// TIA Portal project "EMS" (V15.1)

(* hardware
DEVICE "HMI_SDC"  TP1500 Comfort
   slot 0: "HMI_SDC"  TP1500 Comfort  6AV2 124-0QC02-0AX1  15.1.0.0
   slot 1: "HMI_RT_2"  TP1500 Comfort  6AV2 124-0QC02-0AX1  15.1.0.0
   slot 5: "HMI_SDC._CP_2"  PROFINET Interface  15.0.1.0
      slot 1: "PROFINET Schnittstelle_1"  PROFINET Interface
         slot 1: "Port_1"  Port
         slot 2: "Port_2"  Port
   slot 6: "HMI_SDC._CP_1"  PROFINET Interface  15.0.1.0
      slot 1: "PROFINET Schnittstelle_GBit"  PROFINET Interface
         slot 1: "Port_1"  Port
   slot 7: "HMI_SDC.I/DP_CP_1"  MPI/DP Interface  15.0.1.0
DEVICE "SCALANCE W client"  SCALANCE W-Station
   slot 0: "SCALANCE W rack"  Rail
   slot 0: "_wlan"  SCALANCE W734-1 RJ45 US  6GK5 734-1FX00-0AB0  V6.2
DEVICE "S71500/ET200MP station_1"  S7-1500 station
   slot 0: "Rail_0"  Rack  6ES7 590-1***0-0AA0
   slot 1: "SDC_PLC"  CPU 1518F-4 PN/DP  6ES7 518-4FP00-0AB0  V2.6
      slot 3: "CPU display_1"  6ES7591-1BA00-0AA0
   slot 2: "DI 16x24VDC BA_1"  DI 16x24VDC BA  6ES7 521-1BH10-0AA0  V1.0
   slot 3: "DQ 16x24VDC/0.5A BA_1"  DQ 16x24VDC/0.5A BA  6ES7 522-1BH10-0AA0  V1.0
DEVICE "ET 200SP station_2"  ET 200SP-Station
   slot 0: "Rack_0"  Rack  6ES5 710-8MAx1
   slot 1: "_PLC"  CPU 1512SP F-1 PN  6ES7 512-1SK01-0AB0  V2.1
   slot 2: "F-DI 8x24VDC HF_1"  F-DI 8x24VDC HF  6ES7 136-6BA00-0CA0  V1.0
      slot 1: "F-DI 8x24VDC HF_1"  F-DI 8x24VDC HF
   slot 3: "F-DQ 4x24VDC/2A PM HF_1"  F-DQ 4x24VDC/2A PM HF  6ES7 136-6DB00-0CA0  V1.0
      slot 1: "F-DQ 4x24VDC/2A PM HF_1"  F-DQ 4x24VDC/2A PM HF
   slot 4: "DI 16x24VDC ST_1"  DI 16x24VDC ST  6ES7 131-6BH00-0BA0  V1.1
      slot 1: "DI 16x24VDC ST_1"  DI 16x24VDC ST
   slot 5: "DQ 8x24VDC/0.5A ST_1"  DQ 8x24VDC/0.5A ST  6ES7 132-6BF01-0BA0  V0.0
      slot 1: "DQ 8x24VDC/0.5A ST_1"  DQ 8x24VDC/0.5A ST
   slot 6: "Server module_1"  Server module  6ES7 193-6PA00-0AA0  V1.1
      slot 1: "Server module_1"  Server module
   slot 127: "BA 2xRJ45"  BA 2xRJ45  6ES7 193-6AR00-0AA0  V0.0
      slot 32769: "Port_1"  6ES7 193-6AR00-0AA0
      slot 32770: "Port_2"  6ES7 193-6AR00-0AA0
DEVICE "GSD device_4"  GSD.Device.PN
   slot 0: "Rack"  Rack  V1.0
   slot 0: "_DRIVE"  SINAMICS G120D CU240D-2 PN(-F) V4.7  6SL3 544-0FB2x-1Fxx  V4.70
      slot 0: "SINAMICS G120D CU240D-2 PN(-F) V4.7"  SINAMICS G120D CU240D-2 PN(-F) V4.7
      slot 1: "PN-IO"  PN-IO
         slot 1: "Port 1"  Port 1
         slot 2: "Port 2"  Port 2
      slot 1: "Drive_1"  Drive
         slot 0: "Module Access Point"  Module Access Point
   slot 2: "SIEMENS telegram 352, PZD-6/6"  SIEMENS telegram 352, PZD-6/6
DEVICE "GSD device_1"  GSD.Device.PN
   slot 0: "Rack"  Rack  V1.0
   slot 0: "_ENCODER"  PCV-F200-B17-6011 Position Encoder  PXVxx-F200-B17-V1D-6011
      slot 0: "PCV-F200-B17-6011 Position Encoder"  PCV-F200-B17-6011 Position Encoder
      slot 1: "Interface"  Interface
         slot 1: "Port 1"  Port 1
         slot 2: "Port 2"  Port 2
      slot 1: "Configuration_1"  Configuration
         slot 0: "Configuration"  Configuration
   slot 2: "status_1"  status
      slot 0: "status"  status
   slot 3: "x position_1"  x position
      slot 0: "x position"  x position
   slot 4: "y position_1"  y position
      slot 0: "y position"  y position
DEVICE "GSD device_6"  GSD.Device.PN
   slot 0: "Rack"  Rack  V1.0
   slot 0: "_HMI"  IRD400  6ES7 292-0AA50-1AA0  R01.00.00
      slot 0: "IRD400"  IRD400
      slot 1: "PNIO"  PNIO
         slot 1: "Port 1"  Port 1
         slot 2: "Port 2"  Port 2
      slot 1: "IR Remote Control_1"  IR Remote Control
         slot 0: "IR Remote Control"  IR Remote Control
      slot 2: "Display and LED _1"  Display and LED 
         slot 0: "Display and LED"  Display and LED 
      slot 3: "DIO_1"  DIO
         slot 0: "DIO"  DIO
      slot 4: "IR-P2P_1"  IR-P2P
         slot 0: "IR-P2P"  IR-P2P
      slot 5: "Device Control_1"  Device Control
         slot 0: "Device Control"  Device Control
DEVICE "SCALANCE W access point"  SCALANCE W-Station
   slot 0: "SCALANCE W rack"  Rail
   slot 0: "WLAN_1"  SCALANCE W788-1 M12 US  6GK5 788-1GD00-0AB0  V6.2
DEVICE "GSD device_11"  GSD.Device.PN
   slot 0: "Rack"  Rack  V1.0
   slot 0: "plx32-pnd"  PLX32-EIP-PND  EPD2  1.02.002
      slot 0: "PLX32-EIP-PND"  PLX32-EIP-PND
      slot 1: "Interface1"  Interface1
         slot 1: "Port1"  Port1
   slot 1: "INPUT 512 Byte_1"  INPUT 512 Byte
      slot 0: "INPUT 512 Byte"  INPUT 512 Byte
   slot 2: "OUTPUT 512 Byte_1"  OUTPUT 512 Byte
      slot 0: "OUTPUT 512 Byte"  OUTPUT 512 Byte
   slot 3: "INPUT 256 Byte_3"  INPUT 256 Byte
      slot 0: "INPUT 256 Byte"  INPUT 256 Byte
   slot 4: "OUTPUT 256 Byte_3"  OUTPUT 256 Byte
      slot 0: "OUTPUT 256 Byte"  OUTPUT 256 Byte
   slot 5: "INPUT 256 Byte_2"  INPUT 256 Byte
      slot 0: "INPUT 256 Byte"  INPUT 256 Byte
   slot 6: "OUTPUT 256 Byte_2"  OUTPUT 256 Byte
      slot 0: "OUTPUT 256 Byte"  OUTPUT 256 Byte
   slot 7: "INPUT 256 Byte_1"  INPUT 256 Byte
      slot 0: "INPUT 256 Byte"  INPUT 256 Byte
   slot 8: "OUTPUT 256 Byte_1"  OUTPUT 256 Byte
      slot 0: "OUTPUT 256 Byte"  OUTPUT 256 Byte
*)

// ===== PLC "SDC_PLC"  CPU 1518F-4 PN/DP =====

VAR_GLOBAL   // PLC tag table "Default tag table"
   "LinePLC1_RD_ready" AT %I4248.0 : Bool;
   "EMS_ProductionSpeedRef" AT %IW6130 : Word;
   "EMS_CarrierSpeedRef" AT %IW6126 : Word;
   "SDC_C2_OUT_W9" AT %QW468 : Word;
   "System_Byte" AT %MB1 : Byte;
   "FirstScan" AT %M1.0 : Bool;
   "DiagStatusUpdate" AT %M1.1 : Bool;
   "AlwaysTRUE" AT %M1.2 : Bool;
   "AlwaysFALSE" AT %M1.3 : Bool;
   "Clock_Byte" AT %MB0 : Byte;
   "Clock_10Hz" AT %M0.0 : Bool;
   "Clock_5Hz" AT %M0.1 : Bool;
   "Clock_2.5Hz" AT %M0.2 : Bool;
   "Clock_2Hz" AT %M0.3 : Bool;
   "Clock_1.25Hz" AT %M0.4 : Bool;
   "Clock_1Hz" AT %M0.5 : Bool;
   "Clock_0.625Hz" AT %M0.6 : Bool;
   "Clock_0.5Hz" AT %M0.7 : Bool;
   "tem" AT %M2.0 : Bool;
   "reset" AT %M2.1 : Bool;
   "ZoneCnt" AT %MW4 : Int;
   "Totalcar" AT %MW6 : Int;
   "Tag_3" AT %M2.2 : Bool;
   "carrierzone" AT %MW8 : Int;
   "Carriercnt" AT %MW10 : Int;
   "Carriercnt(1)" AT %MW12 : Int;
   "carrposn" AT %MW14 : Int;
   "IndexArraytemp" AT %MW20 : Int;
   "tempsort" AT %M2.4 : Bool;
   "tempenable2" AT %M2.5 : Bool;
   "tempenable3" AT %M2.6 : Bool;
   "tempenable4" AT %M2.7 : Bool;
   "tempenable5" AT %M3.0 : Bool;
   "tempenable7" AT %M3.1 : Bool;
   "tempblock" AT %M3.2 : Bool;
   "CarrierCounterGbl" AT %MW16 : Int;
   "temp" AT %M3.3 : Bool;
   "cARRIERTESTPOINT" AT %MW18 : Int;
   "cARRIERTESTPOINTBOOL" AT %M3.4 : Bool;
   "cARIERLOOPCOUNT" AT %MW22 : Int;
   "cARIERLOOPCOUNT2" AT %MW24 : Int;
   "tempcarrier27cmdfwd" AT %MW26 : Int;
   "tempcarrier27cmdfwd1" AT %M3.5 : Bool;
   "ZoneCounterGbl" AT %MW28 : Int;
   "IndiconTempDebugON" AT %M3.6 : Bool;
   "HMI_EMS_Nr" AT %MW30 : Int;
   "HMI_EMS_Nr_Calc1" AT %MW32 : Int;
   "HMI_EMS_Nr_Calc2" AT %MW34 : Int;
   "HMI_EMS_Nr__Flt_Out" AT %MW36 : Int;
   "HMI_EMS_Nr__Warn_Out" AT %MW38 : Int;
   "TrafficCopZoneArrayPosCounter" AT %MW40 : Int;
   "SectionComment" AT %M42.0 : Bool;
   "DuplicateCarrierfound" AT %M42.1 : Bool;
   "FaultReset" AT %M42.2 : Bool;
   "DuplicateCarrierNumber" AT %MW44 : Word;
   "CarrierNumberLoop" AT %MW46 : Int;
   "Zone5_ClearToEnter" AT %M42.3 : Bool;
   "PrevCarrierInTransitMem" AT %M42.4 : Bool;
   "SecondDuplicateCarrierPosition" AT %MW50 : Word;
   "FirstDuplicateCarrierPosition" AT %MW48 : Word;
   "EMS_Fault_Reset" AT %M42.5 : Bool;
   "TCCarrierCounterGbl" AT %MW100 : Int;
   "FC206CarrierLoop" AT %MW52 : Int;
   "FC206PositionLoop" AT %MW54 : Int;
   "CARRIER01_POSITION_SDC_OUT" AT %ID402 : DWord;
   "Temp_Int" AT %MW56 : Int;
   "CARRIER #01   1 STATUS [0].5" AT %M80.5 : Bool;
   "CARRIER #01   CURRENT" AT %MW72 : Int;
   "CARRIER #01   G120D CONTROL WORD.0" AT %M74.0 : Bool;
   "CARRIER #01   G120D CONTROL WORD.1" AT %M74.1 : Bool;
   "CARRIER #01   G120D CONTROL WORD.10" AT %M75.2 : Bool;
   "CARRIER #01   G120D CONTROL WORD.11" AT %M75.3 : Bool;
   "CARRIER #01   G120D CONTROL WORD.12" AT %M75.4 : Bool;
   "CARRIER #01   G120D CONTROL WORD.13" AT %M75.5 : Bool;
   "CARRIER #01   G120D CONTROL WORD.14" AT %M75.6 : Bool;
   "CARRIER #01   G120D CONTROL WORD.15" AT %M75.7 : Bool;
   "CARRIER #01   G120D CONTROL WORD.2" AT %M74.2 : Bool;
   "CARRIER #01   G120D CONTROL WORD.3" AT %M74.3 : Bool;
   "CARRIER #01   G120D CONTROL WORD.4" AT %M74.4 : Bool;
   "CARRIER #01   G120D CONTROL WORD.5" AT %M74.5 : Bool;
   "CARRIER #01   G120D CONTROL WORD.6" AT %M74.6 : Bool;
   "CARRIER #01   G120D CONTROL WORD.7" AT %M74.7 : Bool;
   "CARRIER #01   G120D CONTROL WORD.8" AT %M75.0 : Bool;
   "CARRIER #01   G120D CONTROL WORD.9" AT %M75.1 : Bool;
   "CARRIER #01   G120D STATUS WORD.0" AT %M76.0 : Bool;
   "CARRIER #01   G120D STATUS WORD.1" AT %M76.1 : Bool;
   "CARRIER #01   G120D STATUS WORD.10" AT %M77.2 : Bool;
   "CARRIER #01   G120D STATUS WORD.11" AT %M77.3 : Bool;
   "CARRIER #01   G120D STATUS WORD.12" AT %M77.4 : Bool;
   "CARRIER #01   G120D STATUS WORD.13" AT %M77.5 : Bool;
   "CARRIER #01   G120D STATUS WORD.14" AT %M77.6 : Bool;
   "CARRIER #01   G120D STATUS WORD.15" AT %M77.7 : Bool;
   "CARRIER #01   G120D STATUS WORD.2" AT %M76.2 : Bool;
   "CARRIER #01   G120D STATUS WORD.3" AT %M76.3 : Bool;
   "CARRIER #01   G120D STATUS WORD.4" AT %M76.4 : Bool;
   "CARRIER #01   G120D STATUS WORD.5" AT %M76.5 : Bool;
   "CARRIER #01   G120D STATUS WORD.6" AT %M76.6 : Bool;
   "CARRIER #01   G120D STATUS WORD.7" AT %M76.7 : Bool;
   "CARRIER #01   G120D STATUS WORD.8" AT %M77.0 : Bool;
   "CARRIER #01   G120D STATUS WORD.9" AT %M77.1 : Bool;
   "CARRIER #01   POSITION" AT %MW78 : Int;
   "CARRIER #01 480VPowerOn_MDCB1" AT %M80.0 : Bool;
   "CARRIER #01 CrashDetectSW" AT %M80.1 : Bool;
   "CARRIER #01 DCsupplyOnPSCB2" AT %M80.2 : Bool;
   "CARRIER #01 FaultLight_LH" AT %M80.3 : Bool;
   "CARRIER #01 FaultLight_RH" AT %M80.4 : Bool;
   "CARRIER #01 PB1_ProdHoldLH" AT %M80.6 : Bool;
   "CARRIER #01 PB2_ResetLH" AT %M80.7 : Bool;
   "CARRIER #01 PB3_ProdHoldRH" AT %M81.0 : Bool;
   "CARRIER #01 PB4_ResetRH" AT %M81.1 : Bool;
   "CARRIER #01 RunLight_LH" AT %M81.2 : Bool;
   "CARRIER #01 RunLight_RH" AT %M81.3 : Bool;
   "CARRIER #01 SitopSelectStatus" AT %M81.4 : Bool;
   "CARRIER #01 SpareInput(2_1)" AT %M81.5 : Bool;
   "CARRIER #01 SpareInput(2_2)" AT %M81.6 : Bool;
   "CARRIER #01 SpareInput(2_3)" AT %M81.7 : Bool;
   "CARRIER #01 SpareInput(2_4)" AT %M82.0 : Bool;
   "CARRIER #01 SpareInput(2_5)" AT %M82.1 : Bool;
   "CARRIER #01 SpareInput(2_6)" AT %M82.2 : Bool;
   "CARRIER #01 SpareInput(2_7)" AT %M82.3 : Bool;
   "CARRIER #01 SpareInput(4_1)" AT %M82.4 : Bool;
   "CARRIER #01 SpareInput(4_14)" AT %M82.5 : Bool;
   "CARRIER #01 SpareInput(4_15)" AT %M82.6 : Bool;
   "CARRIER #01 SpareInput(4_16)" AT %M82.7 : Bool;
   "CARRIER #01 SpareInput(4_17)" AT %M83.0 : Bool;
   "CARRIER #01 SpareInput(4_2)" AT %M83.1 : Bool;
   "CARRIER #01 SpareInput(4_5)" AT %M83.2 : Bool;
   "CARRIER #01 SpareInput(4_6)" AT %M83.3 : Bool;
   "CARRIER #01 SpareInput(4_7)" AT %M83.4 : Bool;
   "CARRIER #01 SpareOutput(5_5)" AT %M83.5 : Bool;
   "CARRIER #01 SpareOutput(5_6)" AT %M83.6 : Bool;
   "CARRIER #01 SpareOutput(5_7)" AT %M83.7 : Bool;
   "CARRIER #01 SpareSafetyOutput(3_1)" AT %M84.0 : Bool;
   "CARRIER #01 SpareSafetyOutput(3_2)" AT %M84.1 : Bool;
   "CARRIER #01 SpareSafetyOutput(3_3)" AT %M84.2 : Bool;
   "CARRIER #01 SpareSafetyOutput(3_4)" AT %M84.3 : Bool;
   "CARRIER #01 SpareSafetyOutput(3_5)" AT %M84.4 : Bool;
   "CARRIER #01 SpareSafetyOutput(3_6)" AT %M84.5 : Bool;
   "CARRIER #01 SpareSafetyOutput(3_7)" AT %M84.6 : Bool;
   "Carrier #01_ At Command Position" AT %M84.7 : Bool;
   "Carrier #01_ Carrier in zone" AT %MW86 : Int;
   "Carrier #01_ Next carrier number" AT %MW88 : Int;
   "Carrier 1  Drive Status" AT %I412.1 : Bool;
   "Carrier 1 HMI Status" AT %I412.2 : Bool;
   "Carrier 1 PnF Encoder Status" AT %I412.0 : Bool;
   "Carrier 1 Profinet Fault" AT %I410.7 : Bool;
   "Carrier 2  Drive Status" AT %I432.1 : Bool;
   "Carrier 2 HMI Status" AT %I432.2 : Bool;
   "Carrier 2 PnF Encoder Status" AT %I432.0 : Bool;
   "Carrier 2 Profinet Fault" AT %I430.7 : Bool;
   "Carrier 3  Drive Status" AT %I452.1 : Bool;
   "Carrier 3 HMI Status" AT %I452.2 : Bool;
   "Carrier 3 PnF Encoder Status" AT %I452.0 : Bool;
   "Carrier 4  Drive Status" AT %I472.1 : Bool;
   "Carrier 4 HMI Status" AT %I472.2 : Bool;
   "Carrier 4 PnF Encoder Status" AT %I472.0 : Bool;
   "Carrier 4 Profinet Fault" AT %I470.7 : Bool;
   "Carrier_Index_HMI" AT %MW70 : Int;
   "HMI_Zone_Nr" AT %MW102 : Int;
END_VAR

VAR_GLOBAL CONSTANT   // PLC tag table "UserDiag_Constants"
   "USERDIAG_IOSYSTEM_1" : Int := 1;   // Index for first IO-System/DP-Mastersystem
   "USERDIAG_IOSYSTEM_2" : Int := 2;   // Index for second IO-System/DP-Mastersystem
   "USERDIAG_DEVICES_PER_SCREEN_UPPER_LIM" : Int := 128;   // Upper limit of devices per HMI screen
   "USERDIAG_SLOTS_PER_SCREEN_UPPER_LIM" : Int := 31;   // Upper limit of slots per HMI screen
   "USERDIAG_SLOTS_PER_DEVICE_UPPER_LIM" : Int := 31;   // max number of modules per device
   "USERDIAG_DEVICES_PER_IO_SYSTEM_UPPER_LIM" : Int := 128;   // Upper limit of devices/slaves per IO-System/DP-Mastersystem
   "USERDIAG_SLOTS_PER_PLC_UPPER_LIM" : Int := 31;   // max number of local modules
   "USERDIAG_IO_SYSTEMS_UPPER_LIM" : Int := 2;   // Upper limit of IO-Systems/DP-Mastersystems
   "USERDIAG_IOSYSTEM_3" : Int := 3;   // Index for third IO-System/DP-Mastersystem
END_VAR

VAR_GLOBAL   // PLC tag table "Carrier_SDC_TagTable"
   "Carrier_01_Status" AT %IW400 : Word;   // CARRIER STATUS WORD
   "Carrier_01_Status.0" AT %I400.0 : Bool;   // HEARTBEAT
   "Carrier_01_Status.1" AT %I400.1 : Bool;   // MANUAL
   "Carrier_01_Status.2" AT %I400.2 : Bool;   // IN_AUTO
   "Carrier_01_Status.3" AT %I400.3 : Bool;   // POSITIONING_COMPLETE
   "Carrier_01_Status.4" AT %I400.4 : Bool;   // PRODUCTION HOLD
   "Carrier_01_Status.5" AT %I400.5 : Bool;   // CARRIER MOVING FORWARD
   "Carrier_01_Status.6" AT %I400.6 : Bool;   // CARRIER MOVING REVERSE
   "Carrier_01_Status.7" AT %I400.7 : Bool;   // CARRIER FAULT
   "Carrier_01_Status.8" AT %I401.0 : Bool;   // CRASH DETECT TRIPPED
   "Carrier_01_Status.9" AT %I401.1 : Bool;
   "Carrier_01_Status.10" AT %I401.2 : Bool;
   "Carrier_01_Status.11" AT %I401.3 : Bool;
   "Carrier_01_Status.12" AT %I401.4 : Bool;
   "Carrier_01_Status.13" AT %I401.5 : Bool;
   "Carrier_01_Status.14" AT %I401.6 : Bool;
   "Carrier_01_Status.15" AT %I401.7 : Bool;
   "Carrier_01_SDCFaultCode" AT %IW402 : Word;   // SDC FAULT CODE
   "Carrier_01_CarrierPosition" AT %ID404 : DWord;   // CARRIER POSITION
   "Carrier_01_CarrierNumber" AT %IW408 : Word;   // CARRIER NUMBER
   "Carrier_01_G120DControlWord" AT %IW410 : Word;   // G120D_STW1_CONTROL
   "Carrier_01_G120DControlWord.0" AT %I410.0 : Bool;   // Bit_00_ON
   "Carrier_01_G120DControlWord.1" AT %I410.1 : Bool;   // Bit_01_AUS2_INH
   "Carrier_01_G120DControlWord.2" AT %I410.2 : Bool;   // Bit_02_AUS3_STOP
   "Carrier_01_G120DControlWord.3" AT %I410.3 : Bool;   // Bit_03_EN
   "Carrier_01_G120DControlWord.4" AT %I410.4 : Bool;   // Bit_04_EN_RAMP
   "Carrier_01_G120DControlWord.5" AT %I410.5 : Bool;   // Bit_05_START_RAMP
   "Carrier_01_G120DControlWord.6" AT %I410.6 : Bool;   // Bit_06_SETPOINT
   "Carrier_01_G120DControlWord.7" AT %I410.7 : Bool;   // Bit_07_RESET
   "Carrier_01_G120DControlWord.8" AT %I411.0 : Bool;   // Bit_08_JOG_R
   "Carrier_01_G120DControlWord.9" AT %I411.1 : Bool;   // Bit_09_JOG_L
   "Carrier_01_G120DControlWord.10" AT %I411.2 : Bool;   // Bit_10_CONTR_PLC
   "Carrier_01_G120DControlWord.11" AT %I411.3 : Bool;   // Bit_11_REVERSE
   "Carrier_01_G120DControlWord.12" AT %I411.4 : Bool;   // Bit_12_BRAKE_RELEASE
   "Carrier_01_G120DControlWord.13" AT %I411.5 : Bool;   // Bit_13_DDS
   "Carrier_01_G120DControlWord.14" AT %I411.6 : Bool;   // Bit_14_DO0
   "Carrier_01_G120DControlWord.15" AT %I411.7 : Bool;   // Bit_15_DO1
   "Carrier_01_G120DStatusWord" AT %IW412 : Word;   // G120D_ZSW1_STATUS
   "Carrier_01_G120DStatusWord.0" AT %I412.0 : Bool;   // Bit_00_READY_RUN
   "Carrier_01_G120DStatusWord.1" AT %I412.1 : Bool;   // Bit_01_READY_ON
   "Carrier_01_G120DStatusWord.2" AT %I412.2 : Bool;   // Bit_02_ENABLE
   "Carrier_01_G120DStatusWord.3" AT %I412.3 : Bool;   // Bit_03_FAULT
   "Carrier_01_G120DStatusWord.4" AT %I412.4 : Bool;   // Bit_04_OFF2
   "Carrier_01_G120DStatusWord.5" AT %I412.5 : Bool;   // Bit_05_OFF3
   "Carrier_01_G120DStatusWord.6" AT %I412.6 : Bool;   // Bit_06_LOCK_OUT
   "Carrier_01_G120DStatusWord.7" AT %I412.7 : Bool;   // Bit_07_WARN
   "Carrier_01_G120DStatusWord.8" AT %I413.0 : Bool;   // Bit_08_NO_DEVIATION
   "Carrier_01_G120DStatusWord.9" AT %I413.1 : Bool;   // Bit_09_CONTR_PLC
   "Carrier_01_G120DStatusWord.10" AT %I413.2 : Bool;   // Bit_10_F_MAX
   "Carrier_01_G120DStatusWord.11" AT %I413.3 : Bool;   // Bit_11_LIMIT_REACHED
   "Carrier_01_G120DStatusWord.12" AT %I413.4 : Bool;   // Bit_12_BRAKE_OPEN
   "Carrier_01_G120DStatusWord.13" AT %I413.5 : Bool;   // Bit_13_NO_OVERTEMP
   "Carrier_01_G120DStatusWord.14" AT %I413.6 : Bool;   // Bit_14_CW_CCW
   "Carrier_01_G120DStatusWord.15" AT %I413.7 : Bool;   // Bit_15_OVERL
   "Carrier_01_Slot2_Input" AT %IW414 : Word;   // SLOT 2 INPUT WORD
   "Carrier_01_CrashDetectSW" AT %I414.0 : Bool;   // CRASH DETECT SW
   "Carrier_01_SpareSafetyInput(2_1)" AT %I414.1 : Bool;   // SPARE SAFETY INPUT
   "Carrier_01_SpareSafetyInput(2_2)" AT %I414.2 : Bool;   // SPARE SAFETY INPUT
   "Carrier_01_SpareSafetyInput(2_3)" AT %I414.3 : Bool;   // SPARE SAFETY INPUT
   "Carrier_01_SpareSafetyInput(2_4)" AT %I414.4 : Bool;   // SPARE SAFETY INPUT
   "Carrier_01_SpareSafetyInput(2_5)" AT %I414.5 : Bool;   // SPARE SAFETY INPUT
   "Carrier_01_SpareSafetyInput(2_6)" AT %I414.6 : Bool;   // SPARE SAFETY INPUT
   "Carrier_01_SpareSafetyInput(2_7)" AT %I414.7 : Bool;   // SPARE SAFETY INPUT
   "Carrier_01_Slot3_SafetyOutput" AT %IW415 : Word;   // SLOT 3 SAFETY OUTPUT WORD
   "Carrier_01_Crash_Detect_OK" AT %I415.0 : Bool;   // CARRIER CRASH DETECT
   "Carrier_01_SpareSafetyOutput(3_1)" AT %I415.1 : Bool;   // SPARE SAFETY OUTPUT
   "Carrier_01_SpareSafetyOutput(3_2)" AT %I415.2 : Bool;   // SPARE SAFETY OUTPUT
   "Carrier_01_SpareSafetyOutput(3_3)" AT %I415.3 : Bool;   // SPARE SAFETY OUTPUT
   "Carrier_01_SpareSafetyOutput(3_4)" AT %I415.4 : Bool;   // SPARE SAFETY OUTPUT
   "Carrier_01_SpareSafetyOutput(3_5)" AT %I415.5 : Bool;   // SPARE SAFETY OUTPUT
   "Carrier_01_SpareSafetyOutput(3_6)" AT %I415.6 : Bool;   // SPARE SAFETY OUTPUT
   "Carrier_01_SpareSafetyOutput(3_7)" AT %I415.7 : Bool;   // SPARE SAFETY OUTPUT
   "Carrier_01_Slot4_Input" AT %IW416 : Word;   // SLOT 4 INPUT WORD
   "Carrier_01_480VPowerOn_MDCB1" AT %I416.0 : Bool;   // 480 VAC POWER ON MDCB 1
   "Carrier_01_SpareInput(4_1)" AT %I416.1 : Bool;   // SPARE INPUT
   "Carrier_01_SpareInput(4_2)" AT %I416.2 : Bool;   // SPARE INPUT
   "Carrier_01_SitopSelectStatus" AT %I416.3 : Bool;   // SITOP SELECT STATUS
   "Carrier_01_DCsupplyOnPSCB2" AT %I416.4 : Bool;   // DC SUPPLY ON PSCB 2
   "Carrier_01_SpareInput(4_5)" AT %I416.5 : Bool;   // SPARE INPUT
   "Carrier_01_SpareInput(4_6)" AT %I416.6 : Bool;   // SPARE INPUT
   "Carrier_01_SpareInput(4_7)" AT %I416.7 : Bool;   // SPARE INPUT
   "Carrier_01_PB1_ProdHoldLH" AT %I417.0 : Bool;   // PB 1 PRODUCTION HOLD LH
   "Carrier_01_PB2_ResetLH" AT %I417.1 : Bool;   // PB 2 RESET LH
   "Carrier_01_PB3_ProdHoldRH" AT %I417.2 : Bool;   // PB 3 PRODUCTION HOLD RH
   "Carrier_01_PB4_ResetRH" AT %I417.3 : Bool;   // PB 4 RESET RH
   "Carrier_01_SpareInput(4_14)" AT %I417.4 : Bool;   // SPARE INPUT
   "Carrier_01_SpareInput(4_15)" AT %I417.5 : Bool;   // SPARE INPUT
   "Carrier_01_SpareInput(4_16)" AT %I417.6 : Bool;   // SPARE INPUT
   "Carrier_01_SpareInput(4_17)" AT %I417.7 : Bool;   // SPARE INPUT
   "Carrier_01_Slot5_Output" AT %IW418 : Word;   // SLOT 5 OUTPUT WORD
   "Carrier_01_IRD400_HMI_24VDC_ENABLE" AT %I418.0 : Bool;   // IRD 400 PANEL HMI 24V DC POWER
   "Carrier_01_FaultLight_LH" AT %I418.1 : Bool;   // FAULT LIGHT LH
   "Carrier_01_RunLight_LH" AT %I418.2 : Bool;   // RUN LIGHT LH
   "Carrier_01_FaultLight_RH" AT %I418.3 : Bool;   // FAULT LIGHT RH
   "Carrier_01_RunLight_RH" AT %I418.4 : Bool;   // RUN LIGHT RH
   "Carrier_01_SpareOutput(5_5)" AT %I418.5 : Bool;   // SPARE OUTPUT
   "Carrier_01_SpareOutput(5_6)" AT %I418.6 : Bool;   // SPARE OUTPUT
   "Carrier_01_SpareOutput(5_7)" AT %I418.7 : Bool;   // SPARE OUTPUT
   "Carrier_01_ActualSpeed" AT %IW420 : Word;   // ACTUAL SPEED
   "Carrier_01_CarrierDriveAlarm" AT %IW422 : Word;   // CARRIER DRIVE ALARM
   "Carrier_01_CarrierDriveWarning" AT %IW424 : Word;   // CARRIER DRIVE WARNING
   "Carrier_02_Status" AT %IW450 : Word;   // CARRIER STATUS WORD
   "Carrier_02_Status.0" AT %I450.0 : Bool;   // HEARTBEAT
   "Carrier_02_Status.1" AT %I450.1 : Bool;   // MANUAL
   "Carrier_02_Status.2" AT %I450.2 : Bool;   // IN_AUTO
   "Carrier_02_Status.3" AT %I450.3 : Bool;   // POSITIONING_COMPLETE
   "Carrier_02_Status.4" AT %I450.4 : Bool;   // PRODUCTION HOLD
   "Carrier_02_Status.5" AT %I450.5 : Bool;   // CARRIER MOVING FORWARD
   "Carrier_02_Status.6" AT %I450.6 : Bool;   // CARRIER MOVING REVERSE
   "Carrier_02_Status.7" AT %I450.7 : Bool;   // CARRIER FAULT
   "Carrier_02_Status.8" AT %I451.0 : Bool;   // CRASH DETECT TRIPPED
   "Carrier_02_Status.9" AT %I451.1 : Bool;
   "Carrier_02_Status.10" AT %I451.2 : Bool;
   "Carrier_02_Status.11" AT %I451.3 : Bool;
   "Carrier_02_Status.12" AT %I451.4 : Bool;
   "Carrier_02_Status.13" AT %I451.5 : Bool;
   "Carrier_02_Status.14" AT %I451.6 : Bool;
   "Carrier_02_Status.15" AT %I451.7 : Bool;
   "Carrier_02_SDCFaultCode" AT %IW452 : Word;   // SDC FAULT CODE
   "Carrier_02_CarrierPosition" AT %ID454 : DWord;   // CARRIER POSITION
   "Carrier_02_CarrierNumber" AT %IW458 : Word;   // CARRIER NUMBER
   "Carrier_02_G120DControlWord" AT %IW460 : Word;   // G120D_STW1_CONTROL
   "Carrier_02_G120DControlWord.0" AT %I460.0 : Bool;   // Bit_00_ON
   "Carrier_02_G120DControlWord.1" AT %I460.1 : Bool;   // Bit_01_AUS2_INH
   "Carrier_02_G120DControlWord.2" AT %I460.2 : Bool;   // Bit_02_AUS3_STOP
   "Carrier_02_G120DControlWord.3" AT %I460.3 : Bool;   // Bit_03_EN
   "Carrier_02_G120DControlWord.4" AT %I460.4 : Bool;   // Bit_04_EN_RAMP
   "Carrier_02_G120DControlWord.5" AT %I460.5 : Bool;   // Bit_05_START_RAMP
   "Carrier_02_G120DControlWord.6" AT %I460.6 : Bool;   // Bit_06_SETPOINT
   "Carrier_02_G120DControlWord.7" AT %I460.7 : Bool;   // Bit_07_RESET
   "Carrier_02_G120DControlWord.8" AT %I461.0 : Bool;   // Bit_08_JOG_R
   "Carrier_02_G120DControlWord.9" AT %I461.1 : Bool;   // Bit_09_JOG_L
   "Carrier_02_G120DControlWord.10" AT %I461.2 : Bool;   // Bit_10_CONTR_PLC
   "Carrier_02_G120DControlWord.11" AT %I461.3 : Bool;   // Bit_11_REVERSE
   "Carrier_02_G120DControlWord.12" AT %I461.4 : Bool;   // Bit_12_BRAKE_RELEASE
   "Carrier_02_G120DControlWord.13" AT %I461.5 : Bool;   // Bit_13_DDS
   "Carrier_02_G120DControlWord.14" AT %I461.6 : Bool;   // Bit_14_DO0
   "Carrier_02_G120DControlWord.15" AT %I461.7 : Bool;   // Bit_15_DO1
   "Carrier_02_G120DStatusWord" AT %IW462 : Word;   // G120D_ZSW1_STATUS
   "Carrier_02_G120DStatusWord.0" AT %I462.0 : Bool;   // Bit_00_READY_RUN
   "Carrier_02_G120DStatusWord.1" AT %I462.1 : Bool;   // Bit_01_READY_ON
   "Carrier_02_G120DStatusWord.2" AT %I462.2 : Bool;   // Bit_02_ENABLE
   "Carrier_02_G120DStatusWord.3" AT %I462.3 : Bool;   // Bit_03_FAULT
   "Carrier_02_G120DStatusWord.4" AT %I462.4 : Bool;   // Bit_04_OFF2
   "Carrier_02_G120DStatusWord.5" AT %I462.5 : Bool;   // Bit_05_OFF3
   "Carrier_02_G120DStatusWord.6" AT %I462.6 : Bool;   // Bit_06_LOCK_OUT
   "Carrier_02_G120DStatusWord.7" AT %I462.7 : Bool;   // Bit_07_WARN
   "Carrier_02_G120DStatusWord.8" AT %I463.0 : Bool;   // Bit_08_NO_DEVIATION
   "Carrier_02_G120DStatusWord.9" AT %I463.1 : Bool;   // Bit_09_CONTR_PLC
   "Carrier_02_G120DStatusWord.10" AT %I463.2 : Bool;   // Bit_10_F_MAX
   "Carrier_02_G120DStatusWord.11" AT %I463.3 : Bool;   // Bit_11_LIMIT_REACHED
   "Carrier_02_G120DStatusWord.12" AT %I463.4 : Bool;   // Bit_12_BRAKE_OPEN
   "Carrier_02_G120DStatusWord.13" AT %I463.5 : Bool;   // Bit_13_NO_OVERTEMP
   "Carrier_02_G120DStatusWord.14" AT %I463.6 : Bool;   // Bit_14_CW_CCW
   "Carrier_02_G120DStatusWord.15" AT %I463.7 : Bool;   // Bit_15_OVERL
   "Carrier_02_Slot2_Input" AT %IW464 : Word;   // SLOT 2 INPUT WORD
   "Carrier_02_CrashDetectSW" AT %I464.0 : Bool;   // CRASH DETECT SW
   "Carrier_02_SpareSafetyInput(2_1)" AT %I464.1 : Bool;   // SPARE SAFETY INPUT
   "Carrier_02_SpareSafetyInput(2_2)" AT %I464.2 : Bool;   // SPARE SAFETY INPUT
   "Carrier_02_SpareSafetyInput(2_3)" AT %I464.3 : Bool;   // SPARE SAFETY INPUT
   "Carrier_02_SpareSafetyInput(2_4)" AT %I464.4 : Bool;   // SPARE SAFETY INPUT
   "Carrier_02_SpareSafetyInput(2_5)" AT %I464.5 : Bool;   // SPARE SAFETY INPUT
   "Carrier_02_SpareSafetyInput(2_6)" AT %I464.6 : Bool;   // SPARE SAFETY INPUT
   "Carrier_02_SpareSafetyInput(2_7)" AT %I464.7 : Bool;   // SPARE SAFETY INPUT
   "Carrier_02_Slot3_SafetyOutput" AT %IW465 : Word;   // SLOT 3 SAFETY OUTPUT WORD
   "Carrier_02_Crash_Detect_OK" AT %I465.0 : Bool;   // CARRIER CRASH DETECT
   "Carrier_02_SpareSafetyOutput(3_1)" AT %I465.1 : Bool;   // SPARE SAFETY OUTPUT
   "Carrier_02_SpareSafetyOutput(3_2)" AT %I465.2 : Bool;   // SPARE SAFETY OUTPUT
   "Carrier_02_SpareSafetyOutput(3_3)" AT %I465.3 : Bool;   // SPARE SAFETY OUTPUT
   "Carrier_02_SpareSafetyOutput(3_4)" AT %I465.4 : Bool;   // SPARE SAFETY OUTPUT
   "Carrier_02_SpareSafetyOutput(3_5)" AT %I465.5 : Bool;   // SPARE SAFETY OUTPUT
   "Carrier_02_SpareSafetyOutput(3_6)" AT %I465.6 : Bool;   // SPARE SAFETY OUTPUT
   "Carrier_02_SpareSafetyOutput(3_7)" AT %I465.7 : Bool;   // SPARE SAFETY OUTPUT
   "Carrier_02_Slot4_Input" AT %IW466 : Word;   // SLOT 4 INPUT WORD
   "Carrier_02_480VPowerOn_MDCB1" AT %I466.0 : Bool;   // 480 VAC POWER ON MDCB 1
   "Carrier_02_SpareInput(4_1)" AT %I466.1 : Bool;   // SPARE INPUT
   "Carrier_02_SpareInput(4_2)" AT %I466.2 : Bool;   // SPARE INPUT
   "Carrier_02_SitopSelectStatus" AT %I466.3 : Bool;   // SITOP SELECT STATUS
   "Carrier_02_DCsupplyOnPSCB2" AT %I466.4 : Bool;   // DC SUPPLY ON PSCB 2
   "Carrier_02_SpareInput(4_5)" AT %I466.5 : Bool;   // SPARE INPUT
   "Carrier_02_SpareInput(4_6)" AT %I466.6 : Bool;   // SPARE INPUT
   "Carrier_02_SpareInput(4_7)" AT %I466.7 : Bool;   // SPARE INPUT
   "Carrier_02_PB1_ProdHoldLH" AT %I467.0 : Bool;   // PB 1 PRODUCTION HOLD LH
   "Carrier_02_PB2_ResetLH" AT %I467.1 : Bool;   // PB 2 RESET LH
   "Carrier_02_PB3_ProdHoldRH" AT %I467.2 : Bool;   // PB 3 PRODUCTION HOLD RH
   "Carrier_02_PB4_ResetRH" AT %I467.3 : Bool;   // PB 4 RESET RH
   "Carrier_02_SpareInput(4_14)" AT %I467.4 : Bool;   // SPARE INPUT
   "Carrier_02_SpareInput(4_15)" AT %I467.5 : Bool;   // SPARE INPUT
   "Carrier_02_SpareInput(4_16)" AT %I467.6 : Bool;   // SPARE INPUT
   "Carrier_02_SpareInput(4_17)" AT %I467.7 : Bool;   // SPARE INPUT
   "Carrier_02_Slot5_Output" AT %IW468 : Word;   // SLOT 5 OUTPUT WORD
   "Carrier_02_IRD400_HMI_24VDC_ENABLE" AT %I468.0 : Bool;   // IRD 400 PANEL HMI 24V DC POWER
   "Carrier_02_FaultLight_LH" AT %I468.1 : Bool;   // FAULT LIGHT LH
   "Carrier_02_RunLight_LH" AT %I468.2 : Bool;   // RUN LIGHT LH
   "Carrier_02_FaultLight_RH" AT %I468.3 : Bool;   // FAULT LIGHT RH
   "Carrier_02_RunLight_RH" AT %I468.4 : Bool;   // RUN LIGHT RH
   "Carrier_02_SpareOutput(5_5)" AT %I468.5 : Bool;   // SPARE OUTPUT
   "Carrier_02_SpareOutput(5_6)" AT %I468.6 : Bool;   // SPARE OUTPUT
   "Carrier_02_SpareOutput(5_7)" AT %I468.7 : Bool;   // SPARE OUTPUT
   "Carrier_02_ActualSpeed" AT %IW470 : Word;   // ACTUAL SPEED
   "Carrier_02_CarrierDriveAlarm" AT %IW472 : Word;   // CARRIER DRIVE ALARM
   "Carrier_02_CarrierDriveWarning" AT %IW474 : Word;   // CARRIER DRIVE WARNING
   "Carrier_03_Status" AT %IW500 : Word;   // CARRIER STATUS WORD
   "Carrier_03_Status.0" AT %I500.0 : Bool;   // HEARTBEAT
   "Carrier_03_Status.1" AT %I500.1 : Bool;   // MANUAL
   "Carrier_03_Status.2" AT %I500.2 : Bool;   // IN_AUTO
   "Carrier_03_Status.3" AT %I500.3 : Bool;   // POSITIONING_COMPLETE
   "Carrier_03_Status.4" AT %I500.4 : Bool;   // PRODUCTION HOLD
   "Carrier_03_Status.5" AT %I500.5 : Bool;   // CARRIER MOVING FORWARD
   "Carrier_03_Status.6" AT %I500.6 : Bool;   // CARRIER MOVING REVERSE
   "Carrier_03_Status.7" AT %I500.7 : Bool;   // CARRIER FAULT
   "Carrier_03_Status.8" AT %I501.0 : Bool;   // CRASH DETECT TRIPPED
   "Carrier_03_Status.9" AT %I501.1 : Bool;
   "Carrier_03_Status.10" AT %I501.2 : Bool;
   "Carrier_03_Status.11" AT %I501.3 : Bool;
   "Carrier_03_Status.12" AT %I501.4 : Bool;
   "Carrier_03_Status.13" AT %I501.5 : Bool;
   "Carrier_03_Status.14" AT %I501.6 : Bool;
   "Carrier_03_Status.15" AT %I501.7 : Bool;
   "Carrier_03_SDCFaultCode" AT %IW502 : Word;   // SDC FAULT CODE
   "Carrier_03_CarrierPosition" AT %ID504 : DWord;   // CARRIER POSITION
   "Carrier_03_CarrierNumber" AT %IW508 : Word;   // CARRIER NUMBER
   "Carrier_03_G120DControlWord" AT %IW510 : Word;   // G120D_STW1_CONTROL
   "Carrier_03_G120DControlWord.0" AT %I510.0 : Bool;   // Bit_00_ON
   "Carrier_03_G120DControlWord.1" AT %I510.1 : Bool;   // Bit_01_AUS2_INH
   "Carrier_03_G120DControlWord.2" AT %I510.2 : Bool;   // Bit_02_AUS3_STOP
   "Carrier_03_G120DControlWord.3" AT %I510.3 : Bool;   // Bit_03_EN
   "Carrier_03_G120DControlWord.4" AT %I510.4 : Bool;   // Bit_04_EN_RAMP
   "Carrier_03_G120DControlWord.5" AT %I510.5 : Bool;   // Bit_05_START_RAMP
   "Carrier_03_G120DControlWord.6" AT %I510.6 : Bool;   // Bit_06_SETPOINT
   "Carrier_03_G120DControlWord.7" AT %I510.7 : Bool;   // Bit_07_RESET
   "Carrier_03_G120DControlWord.8" AT %I511.0 : Bool;   // Bit_08_JOG_R
   "Carrier_03_G120DControlWord.9" AT %I511.1 : Bool;   // Bit_09_JOG_L
   "Carrier_03_G120DControlWord.10" AT %I511.2 : Bool;   // Bit_10_CONTR_PLC
   "Carrier_03_G120DControlWord.11" AT %I511.3 : Bool;   // Bit_11_REVERSE
   "Carrier_03_G120DControlWord.12" AT %I511.4 : Bool;   // Bit_12_BRAKE_RELEASE
   "Carrier_03_G120DControlWord.13" AT %I511.5 : Bool;   // Bit_13_DDS
   "Carrier_03_G120DControlWord.14" AT %I511.6 : Bool;   // Bit_14_DO0
   "Carrier_03_G120DControlWord.15" AT %I511.7 : Bool;   // Bit_15_DO1
   "Carrier_03_G120DStatusWord" AT %IW512 : Word;   // G120D_ZSW1_STATUS
   "Carrier_03_G120DStatusWord.0" AT %I512.0 : Bool;   // Bit_00_READY_RUN
   "Carrier_03_G120DStatusWord.1" AT %I512.1 : Bool;   // Bit_01_READY_ON
   "Carrier_03_G120DStatusWord.2" AT %I512.2 : Bool;   // Bit_02_ENABLE
   "Carrier_03_G120DStatusWord.3" AT %I512.3 : Bool;   // Bit_03_FAULT
   "Carrier_03_G120DStatusWord.4" AT %I512.4 : Bool;   // Bit_04_OFF2
   "Carrier_03_G120DStatusWord.5" AT %I512.5 : Bool;   // Bit_05_OFF3
   "Carrier_03_G120DStatusWord.6" AT %I512.6 : Bool;   // Bit_06_LOCK_OUT
   "Carrier_03_G120DStatusWord.7" AT %I512.7 : Bool;   // Bit_07_WARN
   "Carrier_03_G120DStatusWord.8" AT %I513.0 : Bool;   // Bit_08_NO_DEVIATION
   "Carrier_03_G120DStatusWord.9" AT %I513.1 : Bool;   // Bit_09_CONTR_PLC
   "Carrier_03_G120DStatusWord.10" AT %I513.2 : Bool;   // Bit_10_F_MAX
   "Carrier_03_G120DStatusWord.11" AT %I513.3 : Bool;   // Bit_11_LIMIT_REACHED
   "Carrier_03_G120DStatusWord.12" AT %I513.4 : Bool;   // Bit_12_BRAKE_OPEN
   "Carrier_03_G120DStatusWord.13" AT %I513.5 : Bool;   // Bit_13_NO_OVERTEMP
   "Carrier_03_G120DStatusWord.14" AT %I513.6 : Bool;   // Bit_14_CW_CCW
   "Carrier_03_G120DStatusWord.15" AT %I513.7 : Bool;   // Bit_15_OVERL
   "Carrier_03_Slot2_Input" AT %IW514 : Word;   // SLOT 2 INPUT WORD
   "Carrier_03_CrashDetectSW" AT %I514.0 : Bool;   // CRASH DETECT SW
   "Carrier_03_SpareSafetyInput(2_1)" AT %I514.1 : Bool;   // SPARE SAFETY INPUT
   "Carrier_03_SpareSafetyInput(2_2)" AT %I514.2 : Bool;   // SPARE SAFETY INPUT
   "Carrier_03_SpareSafetyInput(2_3)" AT %I514.3 : Bool;   // SPARE SAFETY INPUT
   "Carrier_03_SpareSafetyInput(2_4)" AT %I514.4 : Bool;   // SPARE SAFETY INPUT
   "Carrier_03_SpareSafetyInput(2_5)" AT %I514.5 : Bool;   // SPARE SAFETY INPUT
   "Carrier_03_SpareSafetyInput(2_6)" AT %I514.6 : Bool;   // SPARE SAFETY INPUT
   "Carrier_03_SpareSafetyInput(2_7)" AT %I514.7 : Bool;   // SPARE SAFETY INPUT
   "Carrier_03_Slot3_SafetyOutput" AT %IW515 : Word;   // SLOT 3 SAFETY OUTPUT WORD
   "Carrier_03_Crash_Detect_OK" AT %I515.0 : Bool;   // CARRIER CRASH DETECT
   "Carrier_03_SpareSafetyOutput(3_1)" AT %I515.1 : Bool;   // SPARE SAFETY OUTPUT
   "Carrier_03_SpareSafetyOutput(3_2)" AT %I515.2 : Bool;   // SPARE SAFETY OUTPUT
   "Carrier_03_SpareSafetyOutput(3_3)" AT %I515.3 : Bool;   // SPARE SAFETY OUTPUT
   "Carrier_03_SpareSafetyOutput(3_4)" AT %I515.4 : Bool;   // SPARE SAFETY OUTPUT
   "Carrier_03_SpareSafetyOutput(3_5)" AT %I515.5 : Bool;   // SPARE SAFETY OUTPUT
   "Carrier_03_SpareSafetyOutput(3_6)" AT %I515.6 : Bool;   // SPARE SAFETY OUTPUT
   "Carrier_03_SpareSafetyOutput(3_7)" AT %I515.7 : Bool;   // SPARE SAFETY OUTPUT
   "Carrier_03_Slot4_Input" AT %IW516 : Word;   // SLOT 4 INPUT WORD
   "Carrier_03_480VPowerOn_MDCB1" AT %I516.0 : Bool;   // 480 VAC POWER ON MDCB 1
   "Carrier_03_SpareInput(4_1)" AT %I516.1 : Bool;   // SPARE INPUT
   "Carrier_03_SpareInput(4_2)" AT %I516.2 : Bool;   // SPARE INPUT